// TIA Portal project "GzyHzy_1500" (V15)

(* hardware
DEVICE "S71500/ET200MP station_1"  S7-1500 station
   slot 0: "导轨_0"  Rack  6ES7 590-1***0-0AA0
   slot 0: "PM 70W 120/230VAC"  PM 70W 120/230VAC  6EP1332-4BA00
   slot 1: "1#DCC"  CPU 1511-1 PN  6ES7 511-1AK02-0AB0  V2.5
      slot 3: "CPU 显示_1"  6ES7591-1AA00-0AA0
   slot 2: "CP 1542-5_1"  CP 1542-5  6GK7 542-5FX00-0XE0  V1.0
   slot 3: "DI 32x24VDC BA_1"  DI 32x24VDC BA  6ES7 521-1BL10-0AA0  V1.0
   slot 4: "DQ 32x24VDC/0.5A BA_1"  DQ 32x24VDC/0.5A BA  6ES7 522-1BL10-0AA0  V1.0
   slot 5: "AI 8xU/I/RTD/TC ST_1"  AI 8xU/I/RTD/TC ST  6ES7 531-7KF00-0AB0  V2.1
   slot 6: "AI 8xU/I/RTD/TC ST_2"  AI 8xU/I/RTD/TC ST  6ES7 531-7KF00-0AB0  V2.1
   slot 7: "AI 8xU/I/RTD/TC ST_3"  AI 8xU/I/RTD/TC ST  6ES7 531-7KF00-0AB0  V2.1
   slot 8: "AI 8xU/I/RTD/TC ST_4"  AI 8xU/I/RTD/TC ST  6ES7 531-7KF00-0AB0  V2.1
   slot 9: "AI 8xU/I/RTD/TC ST_5"  AI 8xU/I/RTD/TC ST  6ES7 531-7KF00-0AB0  V2.1
   slot 10: "AQ 8xU/I HS_1"  AQ 8xU/I HS  6ES7 532-5HF00-0AB0  V2.1
DEVICE "GSD device_1"  GSD.Device
   slot 0: "机架_0"  Rail
   slot 0: "1#DCC_485"  PB-B-MODBUS  V2.0
DEVICE "S71500/ET200MP station_2"  S7-1500 station
   slot 0: "导轨_0"  Rack  6ES7 590-1***0-0AA0
   slot 0: "PM 70W 120/230VAC"  PM 70W 120/230VAC  6EP1332-4BA00
   slot 1: "1#GZY"  CPU 1511-1 PN  6ES7 511-1AK02-0AB0  V2.5
      slot 3: "CPU 显示_1"  6ES7591-1AA00-0AA0
   slot 2: "CP 1542-5_1"  CP 1542-5  6GK7 542-5FX00-0XE0  V1.0
   slot 3: "DI 32x24VDC BA_1"  DI 32x24VDC BA  6ES7 521-1BL10-0AA0  V1.0
   slot 4: "DI 32x24VDC BA_2"  DI 32x24VDC BA  6ES7 521-1BL10-0AA0  V1.0
   slot 5: "DI 32x24VDC BA_3"  DI 32x24VDC BA  6ES7 521-1BL10-0AA0  V1.0
   slot 6: "DQ 32x24VDC/0.5A BA_1"  DQ 32x24VDC/0.5A BA  6ES7 522-1BL10-0AA0  V1.0
   slot 7: "AI 8xU/I/RTD/TC ST_1"  AI 8xU/I/RTD/TC ST  6ES7 531-7KF00-0AB0  V2.1
   slot 8: "AI 8xU/I/RTD/TC ST_2"  AI 8xU/I/RTD/TC ST  6ES7 531-7KF00-0AB0  V2.1
   slot 9: "AI 8xU/I/RTD/TC ST_3"  AI 8xU/I/RTD/TC ST  6ES7 531-7KF00-0AB0  V2.1
   slot 10: "AI 8xU/I/RTD/TC ST_4"  AI 8xU/I/RTD/TC ST  6ES7 531-7KF00-0AB0  V2.1
   slot 11: "AQ 8xU/I HS_1"  AQ 8xU/I HS  6ES7 532-5HF00-0AB0  V2.1
DEVICE "S71500/ET200MP station_3"  S7-1500 station
   slot 0: "导轨_0"  Rack  6ES7 590-1***0-0AA0
   slot 0: "PM 70W 120/230VAC"  PM 70W 120/230VAC  6EP1332-4BA00
   slot 1: "1#HZY"  CPU 1511-1 PN  6ES7 511-1AK02-0AB0  V2.5
      slot 3: "CPU 显示_1"  6ES7591-1AA00-0AA0
   slot 2: "CP 1542-5_1"  CP 1542-5  6GK7 542-5FX00-0XE0  V1.0
   slot 3: "DI 32x24VDC BA_1"  DI 32x24VDC BA  6ES7 521-1BL10-0AA0  V1.0
   slot 4: "DI 32x24VDC BA_2"  DI 32x24VDC BA  6ES7 521-1BL10-0AA0  V1.0
   slot 5: "DQ 32x24VDC/0.5A BA_1"  DQ 32x24VDC/0.5A BA  6ES7 522-1BL10-0AA0  V1.0
   slot 6: "AI 8xU/I/RTD/TC ST_1"  AI 8xU/I/RTD/TC ST  6ES7 531-7KF00-0AB0  V2.1
   slot 7: "AI 8xU/I/RTD/TC ST_2"  AI 8xU/I/RTD/TC ST  6ES7 531-7KF00-0AB0  V2.1
   slot 8: "AQ 8xU/I HS_1"  AQ 8xU/I HS  6ES7 532-5HF00-0AB0  V2.1
DEVICE "S71500/ET200MP station_4"  S7-1500 station
   slot 0: "导轨_0"  Rack  6ES7 590-1***0-0AA0
   slot 2: "1#HZY_YTZ"  IM 155-5 DP ST  6ES7 155-5BA00-0AB0  V3.0
   slot 3: "DI 16x24VDC BA_1"  DI 16x24VDC BA  6ES7 521-1BH10-0AA0  V1.0
   slot 4: "DI 16x24VDC BA_2"  DI 16x24VDC BA  6ES7 521-1BH10-0AA0  V1.0
   slot 5: "DQ 16x24VDC/0.5A BA_1"  DQ 16x24VDC/0.5A BA  6ES7 522-1BH10-0AA0  V1.0
   slot 6: "AI 8xU/I/RTD/TC ST_1"  AI 8xU/I/RTD/TC ST  6ES7 531-7KF00-0AB0  V2.1
   slot 7: "AI 8xU/I/RTD/TC ST_2"  AI 8xU/I/RTD/TC ST  6ES7 531-7KF00-0AB0  V2.1
   slot 8: "AI 8xU/I/RTD/TC ST_3"  AI 8xU/I/RTD/TC ST  6ES7 531-7KF00-0AB0  V2.1
   slot 9: "AQ 8xU/I HS_1"  AQ 8xU/I HS  6ES7 532-5HF00-0AB0  V2.1
   slot 10: "DI 32x24VDC BA_1"  DI 32x24VDC BA  6ES7 521-1BL10-0AA0  V1.0
   slot 11: "AI 8xU/I/RTD/TC ST_4"  AI 8xU/I/RTD/TC ST  6ES7 531-7KF00-0AB0  V2.1
   slot 12: "AQ 8xU/I HS_2"  AQ 8xU/I HS  6ES7 532-5HF00-0AB0  V2.1
DEVICE "S71500/ET200MP station_5"  S7-1500 station
   slot 0: "导轨_0"  Rack  6ES7 590-1***0-0AA0
   slot 2: "1#HZY_PLZ"  IM 155-5 DP ST  6ES7 155-5BA00-0AB0  V3.0
   slot 3: "DI 16x24VDC BA_1"  DI 16x24VDC BA  6ES7 521-1BH10-0AA0  V1.0
   slot 4: "DI 16x24VDC BA_2"  DI 16x24VDC BA  6ES7 521-1BH10-0AA0  V1.0
   slot 5: "DI 16x24VDC BA_3"  DI 16x24VDC BA  6ES7 521-1BH10-0AA0  V1.0
   slot 6: "DQ 16x24VDC/0.5A BA_1"  DQ 16x24VDC/0.5A BA  6ES7 522-1BH10-0AA0  V1.0
   slot 7: "AI 8xU/I/RTD/TC ST_3"  AI 8xU/I/RTD/TC ST  6ES7 531-7KF00-0AB0  V2.1
   slot 8: "AQ 8xU/I HS_1"  AQ 8xU/I HS  6ES7 532-5HF00-0AB0  V2.1
DEVICE "GSD device_2"  GSD.Device
   slot 0: "机架_0"  Rail
   slot 0: "1#HZY_485"  PB-B-MODBUS  V2.0
DEVICE "GSD device_5"  GSD.Device
   slot 0: "机架_0"  Rail
   slot 0: "1#GZY_485"  PB-B-MODBUS  V2.0
DEVICE "S71500/ET200MP station_6"  S7-1500 station
   slot 0: "导轨_0"  Rack  6ES7 590-1***0-0AA0
   slot 0: "PM 70W 120/230VAC"  PM 70W 120/230VAC  6EP1332-4BA00
   slot 1: "2#DCC"  CPU 1511-1 PN  6ES7 511-1AK02-0AB0  V2.5
      slot 3: "CPU 显示_1"  6ES7591-1AA00-0AA0
   slot 2: "CP 1542-5_1"  CP 1542-5  6GK7 542-5FX00-0XE0  V1.0
   slot 3: "DI 32x24VDC BA_1"  DI 32x24VDC BA  6ES7 521-1BL10-0AA0  V1.0
   slot 4: "DQ 32x24VDC/0.5A BA_1"  DQ 32x24VDC/0.5A BA  6ES7 522-1BL10-0AA0  V1.0
   slot 5: "AI 8xU/I/RTD/TC ST_1"  AI 8xU/I/RTD/TC ST  6ES7 531-7KF00-0AB0  V2.1
   slot 6: "AI 8xU/I/RTD/TC ST_2"  AI 8xU/I/RTD/TC ST  6ES7 531-7KF00-0AB0  V2.1
   slot 7: "AI 8xU/I/RTD/TC ST_3"  AI 8xU/I/RTD/TC ST  6ES7 531-7KF00-0AB0  V2.1
   slot 8: "AI 8xU/I/RTD/TC ST_4"  AI 8xU/I/RTD/TC ST  6ES7 531-7KF00-0AB0  V2.1
   slot 9: "AI 8xU/I/RTD/TC ST_5"  AI 8xU/I/RTD/TC ST  6ES7 531-7KF00-0AB0  V2.1
   slot 10: "AQ 8xU/I HS_1"  AQ 8xU/I HS  6ES7 532-5HF00-0AB0  V2.1
DEVICE "GSD device_6"  GSD.Device
   slot 0: "机架_0"  Rail
   slot 0: "2#DCC_485"  PB-B-MODBUS  V2.0
DEVICE "S71500/ET200MP station_7"  S7-1500 station
   slot 0: "导轨_0"  Rack  6ES7 590-1***0-0AA0
   slot 0: "PM 70W 120/230VAC"  PM 70W 120/230VAC  6EP1332-4BA00
   slot 1: "2#GZY"  CPU 1511-1 PN  6ES7 511-1AK02-0AB0  V2.5
      slot 3: "CPU 显示_1"  6ES7591-1AA00-0AA0
   slot 2: "CP 1542-5_1"  CP 1542-5  6GK7 542-5FX00-0XE0  V1.0
   slot 3: "DI 32x24VDC BA_1"  DI 32x24VDC BA  6ES7 521-1BL10-0AA0  V1.0
   slot 4: "DI 32x24VDC BA_2"  DI 32x24VDC BA  6ES7 521-1BL10-0AA0  V1.0
   slot 5: "DI 32x24VDC BA_3"  DI 32x24VDC BA  6ES7 521-1BL10-0AA0  V1.0
   slot 6: "DQ 32x24VDC/0.5A BA_1"  DQ 32x24VDC/0.5A BA  6ES7 522-1BL10-0AA0  V1.0
   slot 7: "AI 8xU/I/RTD/TC ST_1"  AI 8xU/I/RTD/TC ST  6ES7 531-7KF00-0AB0  V2.1
   slot 8: "AI 8xU/I/RTD/TC ST_2"  AI 8xU/I/RTD/TC ST  6ES7 531-7KF00-0AB0  V2.1
   slot 9: "AI 8xU/I/RTD/TC ST_3"  AI 8xU/I/RTD/TC ST  6ES7 531-7KF00-0AB0  V2.1
   slot 10: "AI 8xU/I/RTD/TC ST_4"  AI 8xU/I/RTD/TC ST  6ES7 531-7KF00-0AB0  V2.1
   slot 11: "AQ 8xU/I HS_1"  AQ 8xU/I HS  6ES7 532-5HF00-0AB0  V2.1
DEVICE "GSD device_7"  GSD.Device
   slot 0: "机架_0"  Rail
   slot 0: "2#GZY_485"  PB-B-MODBUS  V2.0
DEVICE "S71500/ET200MP station_8"  S7-1500 station
   slot 0: "导轨_0"  Rack  6ES7 590-1***0-0AA0
   slot 0: "PM 70W 120/230VAC"  PM 70W 120/230VAC  6EP1332-4BA00
   slot 1: "2#HZY"  CPU 1511-1 PN  6ES7 511-1AK02-0AB0  V2.5
      slot 3: "CPU 显示_1"  6ES7591-1AA00-0AA0
   slot 2: "CP 1542-5_1"  CP 1542-5  6GK7 542-5FX00-0XE0  V1.0
   slot 3: "DI 32x24VDC BA_1"  DI 32x24VDC BA  6ES7 521-1BL10-0AA0  V1.0
   slot 4: "DI 32x24VDC BA_2"  DI 32x24VDC BA  6ES7 521-1BL10-0AA0  V1.0
   slot 5: "DQ 32x24VDC/0.5A BA_1"  DQ 32x24VDC/0.5A BA  6ES7 522-1BL10-0AA0  V1.0
   slot 6: "AI 8xU/I/RTD/TC ST_1"  AI 8xU/I/RTD/TC ST  6ES7 531-7KF00-0AB0  V2.1
   slot 7: "AI 8xU/I/RTD/TC ST_2"  AI 8xU/I/RTD/TC ST  6ES7 531-7KF00-0AB0  V2.1
   slot 8: "AQ 8xU/I HS_1"  AQ 8xU/I HS  6ES7 532-5HF00-0AB0  V2.1
DEVICE "S71500/ET200MP station_9"  S7-1500 station
   slot 0: "导轨_0"  Rack  6ES7 590-1***0-0AA0
   slot 2: "2#HZY_YTZ"  IM 155-5 DP ST  6ES7 155-5BA00-0AB0  V3.0
   slot 3: "DI 16x24VDC BA_1"  DI 16x24VDC BA  6ES7 521-1BH10-0AA0  V1.0
   slot 4: "DI 16x24VDC BA_2"  DI 16x24VDC BA  6ES7 521-1BH10-0AA0  V1.0
   slot 5: "DQ 16x24VDC/0.5A BA_1"  DQ 16x24VDC/0.5A BA  6ES7 522-1BH10-0AA0  V1.0
   slot 6: "AI 8xU/I/RTD/TC ST_1"  AI 8xU/I/RTD/TC ST  6ES7 531-7KF00-0AB0  V2.1
   slot 7: "AI 8xU/I/RTD/TC ST_2"  AI 8xU/I/RTD/TC ST  6ES7 531-7KF00-0AB0  V2.1
   slot 8: "AI 8xU/I/RTD/TC ST_3"  AI 8xU/I/RTD/TC ST  6ES7 531-7KF00-0AB0  V2.1
   slot 9: "AQ 8xU/I HS_1"  AQ 8xU/I HS  6ES7 532-5HF00-0AB0  V2.1
   slot 10: "DI 32x24VDC BA_1"  DI 32x24VDC BA  6ES7 521-1BL10-0AA0  V1.0
   slot 11: "AI 8xU/I/RTD/TC ST_4"  AI 8xU/I/RTD/TC ST  6ES7 531-7KF00-0AB0  V2.1
   slot 12: "AQ 8xU/I HS_2"  AQ 8xU/I HS  6ES7 532-5HF00-0AB0  V2.1
DEVICE "S71500/ET200MP station_10"  S7-1500 station
   slot 0: "导轨_0"  Rack  6ES7 590-1***0-0AA0
   slot 2: "2#HZY_PLZ"  IM 155-5 DP ST  6ES7 155-5BA00-0AB0  V3.0
   slot 3: "DI 16x24VDC BA_1"  DI 16x24VDC BA  6ES7 521-1BH10-0AA0  V1.0
   slot 4: "DI 16x24VDC BA_2"  DI 16x24VDC BA  6ES7 521-1BH10-0AA0  V1.0
   slot 5: "DI 16x24VDC BA_3"  DI 16x24VDC BA  6ES7 521-1BH10-0AA0  V1.0
   slot 6: "DQ 16x24VDC/0.5A BA_1"  DQ 16x24VDC/0.5A BA  6ES7 522-1BH10-0AA0  V1.0
   slot 7: "AI 8xU/I/RTD/TC ST_3"  AI 8xU/I/RTD/TC ST  6ES7 531-7KF00-0AB0  V2.1
   slot 8: "AQ 8xU/I HS_1"  AQ 8xU/I HS  6ES7 532-5HF00-0AB0  V2.1
DEVICE "GSD device_8"  GSD.Device
   slot 0: "机架_0"  Rail
   slot 0: "2#HZY_485"  PB-B-MODBUS  V2.0
DEVICE "S71500/ET200MP station_11"  S7-1500 station
   slot 0: "导轨_0"  Rack  6ES7 590-1***0-0AA0
   slot 0: "PM 70W 120/230VAC"  PM 70W 120/230VAC  6EP1332-4BA00
   slot 1: "3#GZY"  CPU 1511-1 PN  6ES7 511-1AK02-0AB0  V2.5
      slot 3: "CPU 显示_1"  6ES7591-1AA00-0AA0
   slot 2: "CP 1542-5_1"  CP 1542-5  6GK7 542-5FX00-0XE0  V1.0
   slot 3: "DI 32x24VDC BA_1"  DI 32x24VDC BA  6ES7 521-1BL10-0AA0  V1.0
   slot 4: "DI 32x24VDC BA_2"  DI 32x24VDC BA  6ES7 521-1BL10-0AA0  V1.0
   slot 5: "DI 32x24VDC BA_3"  DI 32x24VDC BA  6ES7 521-1BL10-0AA0  V1.0
   slot 6: "DQ 32x24VDC/0.5A BA_1"  DQ 32x24VDC/0.5A BA  6ES7 522-1BL10-0AA0  V1.0
   slot 7: "AI 8xU/I/RTD/TC ST_1"  AI 8xU/I/RTD/TC ST  6ES7 531-7KF00-0AB0  V2.1
   slot 8: "AI 8xU/I/RTD/TC ST_2"  AI 8xU/I/RTD/TC ST  6ES7 531-7KF00-0AB0  V2.1
   slot 9: "AI 8xU/I/RTD/TC ST_3"  AI 8xU/I/RTD/TC ST  6ES7 531-7KF00-0AB0  V2.1
   slot 10: "AI 8xU/I/RTD/TC ST_4"  AI 8xU/I/RTD/TC ST  6ES7 531-7KF00-0AB0  V2.1
   slot 11: "AQ 8xU/I HS_1"  AQ 8xU/I HS  6ES7 532-5HF00-0AB0  V2.1
DEVICE "GSD device_11"  GSD.Device
   slot 0: "机架_0"  Rail
   slot 0: "3#GZY_485"  PB-B-MODBUS  V2.0
DEVICE "S71500/ET200MP station_12"  S7-1500 station
   slot 0: "导轨_0"  Rack  6ES7 590-1***0-0AA0
   slot 0: "PM 70W 120/230VAC"  PM 70W 120/230VAC  6EP1332-4BA00
   slot 1: "3#HZY"  CPU 1511-1 PN  6ES7 511-1AK02-0AB0  V2.5
      slot 3: "CPU 显示_1"  6ES7591-1AA00-0AA0
   slot 2: "CP 1542-5_1"  CP 1542-5  6GK7 542-5FX00-0XE0  V1.0
   slot 3: "DI 32x24VDC BA_1"  DI 32x24VDC BA  6ES7 521-1BL10-0AA0  V1.0
   slot 4: "DI 32x24VDC BA_2"  DI 32x24VDC BA  6ES7 521-1BL10-0AA0  V1.0
   slot 5: "DQ 32x24VDC/0.5A BA_1"  DQ 32x24VDC/0.5A BA  6ES7 522-1BL10-0AA0  V1.0
   slot 6: "AI 8xU/I/RTD/TC ST_1"  AI 8xU/I/RTD/TC ST  6ES7 531-7KF00-0AB0  V2.1
   slot 7: "AI 8xU/I/RTD/TC ST_2"  AI 8xU/I/RTD/TC ST  6ES7 531-7KF00-0AB0  V2.1
   slot 8: "AQ 8xU/I HS_1"  AQ 8xU/I HS  6ES7 532-5HF00-0AB0  V2.1
DEVICE "S71500/ET200MP station_14"  S7-1500 station
   slot 0: "导轨_0"  Rack  6ES7 590-1***0-0AA0
   slot 2: "3#HZY_YTZ"  IM 155-5 DP ST  6ES7 155-5BA00-0AB0  V3.0
   slot 3: "DI 16x24VDC BA_1"  DI 16x24VDC BA  6ES7 521-1BH10-0AA0  V1.0
   slot 4: "DI 16x24VDC BA_2"  DI 16x24VDC BA  6ES7 521-1BH10-0AA0  V1.0
   slot 5: "DQ 16x24VDC/0.5A BA_1"  DQ 16x24VDC/0.5A BA  6ES7 522-1BH10-0AA0  V1.0
   slot 6: "AI 8xU/I/RTD/TC ST_1"  AI 8xU/I/RTD/TC ST  6ES7 531-7KF00-0AB0  V2.1
   slot 7: "AI 8xU/I/RTD/TC ST_2"  AI 8xU/I/RTD/TC ST  6ES7 531-7KF00-0AB0  V2.1
   slot 8: "AI 8xU/I/RTD/TC ST_3"  AI 8xU/I/RTD/TC ST  6ES7 531-7KF00-0AB0  V2.1
   slot 9: "AQ 8xU/I HS_1"  AQ 8xU/I HS  6ES7 532-5HF00-0AB0  V2.1
   slot 10: "DI 32x24VDC BA_1"  DI 32x24VDC BA  6ES7 521-1BL10-0AA0  V1.0
   slot 11: "AI 8xU/I/RTD/TC ST_4"  AI 8xU/I/RTD/TC ST  6ES7 531-7KF00-0AB0  V2.1
   slot 12: "AQ 8xU/I HS_2"  AQ 8xU/I HS  6ES7 532-5HF00-0AB0  V2.1
DEVICE "S71500/ET200MP station_13"  S7-1500 station
   slot 0: "导轨_0"  Rack  6ES7 590-1***0-0AA0
   slot 2: "3#HZY_PLZ"  IM 155-5 DP ST  6ES7 155-5BA00-0AB0  V3.0
   slot 3: "DI 16x24VDC BA_1"  DI 16x24VDC BA  6ES7 521-1BH10-0AA0  V1.0
   slot 4: "DI 16x24VDC BA_2"  DI 16x24VDC BA  6ES7 521-1BH10-0AA0  V1.0
   slot 5: "DI 16x24VDC BA_3"  DI 16x24VDC BA  6ES7 521-1BH10-0AA0  V1.0
   slot 6: "DQ 16x24VDC/0.5A BA_1"  DQ 16x24VDC/0.5A BA  6ES7 522-1BH10-0AA0  V1.0
   slot 7: "AI 8xU/I/RTD/TC ST_3"  AI 8xU/I/RTD/TC ST  6ES7 531-7KF00-0AB0  V2.1
   slot 8: "AQ 8xU/I HS_1"  AQ 8xU/I HS  6ES7 532-5HF00-0AB0  V2.1
DEVICE "GSD device_12"  GSD.Device
   slot 0: "机架_0"  Rail
   slot 0: "3#HZY_485"  PB-B-MODBUS  V2.0
DEVICE "S71500/ET200MP station_15"  S7-1500 station
   slot 0: "导轨_0"  Rack  6ES7 590-1***0-0AA0
   slot 0: "PM 70W 120/230VAC"  PM 70W 120/230VAC  6EP1332-4BA00
   slot 1: "4#GZY"  CPU 1511-1 PN  6ES7 511-1AK02-0AB0  V2.5
      slot 3: "CPU 显示_1"  6ES7591-1AA00-0AA0
   slot 2: "CP 1542-5_1"  CP 1542-5  6GK7 542-5FX00-0XE0  V1.0
   slot 3: "DI 32x24VDC BA_1"  DI 32x24VDC BA  6ES7 521-1BL10-0AA0  V1.0
   slot 4: "DI 32x24VDC BA_2"  DI 32x24VDC BA  6ES7 521-1BL10-0AA0  V1.0
   slot 5: "DI 32x24VDC BA_3"  DI 32x24VDC BA  6ES7 521-1BL10-0AA0  V1.0
   slot 6: "DQ 32x24VDC/0.5A BA_1"  DQ 32x24VDC/0.5A BA  6ES7 522-1BL10-0AA0  V1.0
   slot 7: "AI 8xU/I/RTD/TC ST_1"  AI 8xU/I/RTD/TC ST  6ES7 531-7KF00-0AB0  V2.1
   slot 8: "AI 8xU/I/RTD/TC ST_2"  AI 8xU/I/RTD/TC ST  6ES7 531-7KF00-0AB0  V2.1
   slot 9: "AI 8xU/I/RTD/TC ST_3"  AI 8xU/I/RTD/TC ST  6ES7 531-7KF00-0AB0  V2.1
   slot 10: "AI 8xU/I/RTD/TC ST_4"  AI 8xU/I/RTD/TC ST  6ES7 531-7KF00-0AB0  V2.1
   slot 11: "AQ 8xU/I HS_1"  AQ 8xU/I HS  6ES7 532-5HF00-0AB0  V2.1
DEVICE "S71500/ET200MP station_16"  S7-1500 station
   slot 0: "导轨_0"  Rack  6ES7 590-1***0-0AA0
   slot 0: "PM 70W 120/230VAC"  PM 70W 120/230VAC  6EP1332-4BA00
   slot 1: "4#HZY"  CPU 1511-1 PN  6ES7 511-1AK02-0AB0  V2.5
      slot 3: "CPU 显示_1"  6ES7591-1AA00-0AA0
   slot 2: "CP 1542-5_1"  CP 1542-5  6GK7 542-5FX00-0XE0  V1.0
   slot 3: "DI 32x24VDC BA_1"  DI 32x24VDC BA  6ES7 521-1BL10-0AA0  V1.0
   slot 4: "DI 32x24VDC BA_2"  DI 32x24VDC BA  6ES7 521-1BL10-0AA0  V1.0
   slot 5: "DQ 32x24VDC/0.5A BA_1"  DQ 32x24VDC/0.5A BA  6ES7 522-1BL10-0AA0  V1.0
   slot 6: "AI 8xU/I/RTD/TC ST_1"  AI 8xU/I/RTD/TC ST  6ES7 531-7KF00-0AB0  V2.1
   slot 7: "AI 8xU/I/RTD/TC ST_2"  AI 8xU/I/RTD/TC ST  6ES7 531-7KF00-0AB0  V2.1
   slot 8: "AQ 8xU/I HS_1"  AQ 8xU/I HS  6ES7 532-5HF00-0AB0  V2.1
DEVICE "S71500/ET200MP station_17"  S7-1500 station
   slot 0: "导轨_0"  Rack  6ES7 590-1***0-0AA0
   slot 2: "4#HZY_YTZ"  IM 155-5 DP ST  6ES7 155-5BA00-0AB0  V3.0
   slot 3: "DI 16x24VDC BA_1"  DI 16x24VDC BA  6ES7 521-1BH10-0AA0  V1.0
   slot 4: "DI 16x24VDC BA_2"  DI 16x24VDC BA  6ES7 521-1BH10-0AA0  V1.0
   slot 5: "DQ 16x24VDC/0.5A BA_1"  DQ 16x24VDC/0.5A BA  6ES7 522-1BH10-0AA0  V1.0
   slot 6: "AI 8xU/I/RTD/TC ST_1"  AI 8xU/I/RTD/TC ST  6ES7 531-7KF00-0AB0  V2.1
   slot 7: "AI 8xU/I/RTD/TC ST_2"  AI 8xU/I/RTD/TC ST  6ES7 531-7KF00-0AB0  V2.1
   slot 8: "AI 8xU/I/RTD/TC ST_3"  AI 8xU/I/RTD/TC ST  6ES7 531-7KF00-0AB0  V2.1
   slot 9: "AQ 8xU/I HS_1"  AQ 8xU/I HS  6ES7 532-5HF00-0AB0  V2.1
   slot 10: "DI 32x24VDC BA_1"  DI 32x24VDC BA  6ES7 521-1BL10-0AA0  V1.0
   slot 11: "AI 8xU/I/RTD/TC ST_4"  AI 8xU/I/RTD/TC ST  6ES7 531-7KF00-0AB0  V2.1
   slot 12: "AQ 8xU/I HS_2"  AQ 8xU/I HS  6ES7 532-5HF00-0AB0  V2.1
DEVICE "S71500/ET200MP station_18"  S7-1500 station
   slot 0: "导轨_0"  Rack  6ES7 590-1***0-0AA0
   slot 2: "4#HZY_PLZ"  IM 155-5 DP ST  6ES7 155-5BA00-0AB0  V3.0
   slot 3: "DI 16x24VDC BA_1"  DI 16x24VDC BA  6ES7 521-1BH10-0AA0  V1.0
   slot 4: "DI 16x24VDC BA_2"  DI 16x24VDC BA  6ES7 521-1BH10-0AA0  V1.0
   slot 5: "DI 16x24VDC BA_3"  DI 16x24VDC BA  6ES7 521-1BH10-0AA0  V1.0
   slot 6: "DQ 16x24VDC/0.5A BA_1"  DQ 16x24VDC/0.5A BA  6ES7 522-1BH10-0AA0  V1.0
   slot 7: "AI 8xU/I/RTD/TC ST_3"  AI 8xU/I/RTD/TC ST  6ES7 531-7KF00-0AB0  V2.1
   slot 8: "AQ 8xU/I HS_1"  AQ 8xU/I HS  6ES7 532-5HF00-0AB0  V2.1
DEVICE "GSD device_16"  GSD.Device
   slot 0: "机架_0"  Rail
   slot 0: "4#HZY_485"  PB-B-MODBUS  V2.0
DEVICE "S71500/ET200MP station_19"  S7-1500 station
   slot 0: "导轨_0"  Rack  6ES7 590-1***0-0AA0
   slot 0: "PM 70W 120/230VAC"  PM 70W 120/230VAC  6EP1332-4BA00
   slot 1: "1#LM"  CPU 1511-1 PN  6ES7 511-1AK02-0AB0  V2.5
      slot 3: "CPU 显示_1"  6ES7591-1AA00-0AA0
   slot 2: "CP 1542-5_1"  CP 1542-5  6GK7 542-5FX00-0XE0  V1.0
   slot 3: "DI 32x24VDC BA_1"  DI 32x24VDC BA  6ES7 521-1BL10-0AA0  V1.0
   slot 4: "DI 32x24VDC BA_2"  DI 32x24VDC BA  6ES7 521-1BL10-0AA0  V1.0
   slot 5: "DI 32x24VDC BA_3"  DI 32x24VDC BA  6ES7 521-1BL10-0AA0  V1.0
   slot 6: "DQ 32x24VDC/0.5A BA_1"  DQ 32x24VDC/0.5A BA  6ES7 522-1BL10-0AA0  V1.0
   slot 7: "AI 8xU/I/RTD/TC ST_1"  AI 8xU/I/RTD/TC ST  6ES7 531-7KF00-0AB0  V2.1
   slot 8: "AI 8xU/I/RTD/TC ST_2"  AI 8xU/I/RTD/TC ST  6ES7 531-7KF00-0AB0  V2.1
   slot 9: "AI 8xU/I/RTD/TC ST_3"  AI 8xU/I/RTD/TC ST  6ES7 531-7KF00-0AB0  V2.1
   slot 10: "AQ 8xU/I HS_1"  AQ 8xU/I HS  6ES7 532-5HF00-0AB0  V2.1
DEVICE "GSD device_19"  GSD.Device
   slot 0: "机架_0"  Rail
   slot 0: "1#LM_485"  PB-B-MODBUS  V2.0
DEVICE "GSD device_15"  GSD.Device
   slot 0: "机架_0"  Rail
   slot 0: "4#GZY_485"  PB-B-MODBUS  V2.0
DEVICE "GSD device_28"  GSD.Device
   slot 0: "机架_0"  Rail
DEVICE "GSD device_25"  GSD.Device
   slot 0: "机架_0"  Rail
DEVICE "GSD device_21"  GSD.Device
   slot 0: "机架_0"  Rail
DEVICE "GSD device_22"  GSD.Device
   slot 0: "机架_0"  Rail
DEVICE "SINAMICS G_4"  Sinamics.Device
   slot 0: "	_0"  Rail  SinamicsG120Rack-V
   slot 2: "电炉料罐车变频_1"  G120 CU240E-2  6SL3244-0BB12-1BA1  4.7.6
   slot 3: "PM240-2 IP20"  PM240-2 IP20  6SL3210-1PE23-3ULx  -
DEVICE "GSD device_23"  GSD.Device
   slot 0: "机架_0"  Rail
DEVICE "GSD device_24"  GSD.Device
   slot 0: "机架_0"  Rail
DEVICE "GSD device_26"  GSD.Device
   slot 0: "机架_0"  Rail
DEVICE "GSD device_3"  GSD.Device
   slot 0: "机架_0"  Rail
DEVICE "GSD device_4"  GSD.Device
   slot 0: "机架_0"  Rail
DEVICE "GSD device_9"  GSD.Device
   slot 0: "机架_0"  Rail
DEVICE "GSD device_10"  GSD.Device
   slot 0: "机架_0"  Rail
DEVICE "GSD device_13"  GSD.Device
   slot 0: "机架_0"  Rail
DEVICE "GSD device_14"  GSD.Device
   slot 0: "机架_0"  Rail
DEVICE "GSD device_17"  GSD.Device
   slot 0: "机架_0"  Rail
DEVICE "GSD device_18"  GSD.Device
   slot 0: "机架_0"  Rail
DEVICE "S71500/ET200MP station_20"  S7-1500 station
   slot 0: "导轨_0"  Rack  6ES7 590-1***0-0AA0
   slot 0: "PM 70W 120/230VAC"  PM 70W 120/230VAC  6EP1332-4BA00
   slot 1: "1#SBF"  CPU 1511-1 PN  6ES7 511-1AK02-0AB0  V2.5
      slot 3: "CPU 显示_1"  6ES7591-1AA00-0AA0
   slot 2: "CP 1542-5_1"  CP 1542-5  6GK7 542-5FX00-0XE0  V1.0
   slot 3: "DI 32x24VDC BA_1"  DI 32x24VDC BA  6ES7 521-1BL10-0AA0  V1.0
   slot 4: "DI 32x24VDC BA_2"  DI 32x24VDC BA  6ES7 521-1BL10-0AA0  V1.0
   slot 5: "DI 32x24VDC BA_3"  DI 32x24VDC BA  6ES7 521-1BL10-0AA0  V1.0
   slot 6: "DI 32x24VDC BA_4"  DI 32x24VDC BA  6ES7 521-1BL10-0AA0  V1.0
   slot 7: "DI 32x24VDC BA_5"  DI 32x24VDC BA  6ES7 521-1BL10-0AA0  V1.0
   slot 8: "DI 32x24VDC BA_6"  DI 32x24VDC BA  6ES7 521-1BL10-0AA0  V1.0
   slot 9: "PS 25W 24VDC_1"  PS 25W 24VDC  6ES7 505-0KA00-0AB0  V1.0
   slot 10: "DQ 32x24VDC/0.5A BA_1"  DQ 32x24VDC/0.5A BA  6ES7 522-1BL10-0AA0  V1.0
   slot 11: "DQ 32x24VDC/0.5A BA_2"  DQ 32x24VDC/0.5A BA  6ES7 522-1BL10-0AA0  V1.0
DEVICE "S71500/ET200MP station_25"  S7-1500 station
   slot 0: "导轨_0"  Rack  6ES7 590-1***0-0AA0
   slot 0: "PM 70W 120/230VAC"  PM 70W 120/230VAC  6EP1332-4BA00
   slot 1: "2#SBF"  CPU 1511-1 PN  6ES7 511-1AK02-0AB0  V2.5
      slot 3: "CPU 显示_1"  6ES7591-1AA00-0AA0
   slot 2: "CP 1542-5_1"  CP 1542-5  6GK7 542-5FX00-0XE0  V1.0
   slot 3: "DI 32x24VDC BA_1"  DI 32x24VDC BA  6ES7 521-1BL10-0AA0  V1.0
   slot 4: "DI 32x24VDC BA_2"  DI 32x24VDC BA  6ES7 521-1BL10-0AA0  V1.0
   slot 5: "DI 32x24VDC BA_3"  DI 32x24VDC BA  6ES7 521-1BL10-0AA0  V1.0
   slot 6: "DI 32x24VDC BA_4"  DI 32x24VDC BA  6ES7 521-1BL10-0AA0  V1.0
   slot 7: "DI 32x24VDC BA_5"  DI 32x24VDC BA  6ES7 521-1BL10-0AA0  V1.0
   slot 8: "DI 32x24VDC BA_6"  DI 32x24VDC BA  6ES7 521-1BL10-0AA0  V1.0
   slot 9: "PS 25W 24VDC_1"  PS 25W 24VDC  6ES7 505-0KA00-0AB0  V1.0
   slot 10: "DQ 32x24VDC/0.5A BA_1"  DQ 32x24VDC/0.5A BA  6ES7 522-1BL10-0AA0  V1.0
   slot 11: "DQ 32x24VDC/0.5A BA_2"  DQ 32x24VDC/0.5A BA  6ES7 522-1BL10-0AA0  V1.0
DEVICE "S71500/ET200MP station_21"  S7-1500 station
   slot 0: "导轨_0"  Rack  6ES7 590-1***0-0AA0
   slot 2: "1#SBF_1"  IM 155-5 DP ST  6ES7 155-5BA00-0AB0  V3.0
   slot 3: "DI 32x24VDC BA_1"  DI 32x24VDC BA  6ES7 521-1BL10-0AA0  V1.0
   slot 4: "DI 32x24VDC BA_2"  DI 32x24VDC BA  6ES7 521-1BL10-0AA0  V1.0
   slot 5: "DI 32x24VDC BA_3"  DI 32x24VDC BA  6ES7 521-1BL10-0AA0  V1.0
   slot 6: "DQ 32x24VDC/0.5A BA_1"  DQ 32x24VDC/0.5A BA  6ES7 522-1BL10-0AA0  V1.0
   slot 7: "DQ 32x24VDC/0.5A BA_2"  DQ 32x24VDC/0.5A BA  6ES7 522-1BL10-0AA0  V1.0
DEVICE "S71500/ET200MP station_22"  S7-1500 station
   slot 0: "导轨_0"  Rack  6ES7 590-1***0-0AA0
   slot 2: "1#SBF_2"  IM 155-5 DP ST  6ES7 155-5BA00-0AB0  V3.0
   slot 3: "AI 8xU/I/RTD/TC ST_1"  AI 8xU/I/RTD/TC ST  6ES7 531-7KF00-0AB0  V2.1
   slot 4: "AI 8xU/I/RTD/TC ST_2"  AI 8xU/I/RTD/TC ST  6ES7 531-7KF00-0AB0  V2.1
   slot 5: "AI 8xU/I/RTD/TC ST_3"  AI 8xU/I/RTD/TC ST  6ES7 531-7KF00-0AB0  V2.1
   slot 6: "AI 8xU/I/RTD/TC ST_4"  AI 8xU/I/RTD/TC ST  6ES7 531-7KF00-0AB0  V2.1
   slot 7: "AI 8xU/I/RTD/TC ST_5"  AI 8xU/I/RTD/TC ST  6ES7 531-7KF00-0AB0  V2.1
   slot 8: "AQ 8xU/I HS_1"  AQ 8xU/I HS  6ES7 532-5HF00-0AB0  V2.1
   slot 9: "AQ 8xU/I HS_2"  AQ 8xU/I HS  6ES7 532-5HF00-0AB0  V2.1
   slot 10: "AQ 8xU/I HS_3"  AQ 8xU/I HS  6ES7 532-5HF00-0AB0  V2.1
DEVICE "S71500/ET200MP station_23"  S7-1500 station
   slot 0: "导轨_0"  Rack  6ES7 590-1***0-0AA0
   slot 2: "1#SBF_3"  IM 155-5 DP ST  6ES7 155-5BA00-0AB0  V3.0
   slot 3: "DI 32x24VDC BA_1"  DI 32x24VDC BA  6ES7 521-1BL10-0AA0  V1.0
   slot 4: "DI 32x24VDC BA_2"  DI 32x24VDC BA  6ES7 521-1BL10-0AA0  V1.0
   slot 5: "DQ 32x24VDC/0.5A BA_1"  DQ 32x24VDC/0.5A BA  6ES7 522-1BL10-0AA0  V1.0
   slot 6: "AI 8xU/I/RTD/TC ST_1"  AI 8xU/I/RTD/TC ST  6ES7 531-7KF00-0AB0  V2.1
   slot 7: "AI 8xU/I/RTD/TC ST_2"  AI 8xU/I/RTD/TC ST  6ES7 531-7KF00-0AB0  V2.1
   slot 8: "AQ 8xU/I HS_1"  AQ 8xU/I HS  6ES7 532-5HF00-0AB0  V2.1
DEVICE "S71500/ET200MP station_24"  S7-1500 station
   slot 0: "导轨_0"  Rack  6ES7 590-1***0-0AA0
   slot 2: "1#SBF_4"  IM 155-5 DP ST  6ES7 155-5BA00-0AB0  V3.0
   slot 3: "DI 32x24VDC BA_1"  DI 32x24VDC BA  6ES7 521-1BL10-0AA0  V1.0
   slot 4: "DI 32x24VDC BA_2"  DI 32x24VDC BA  6ES7 521-1BL10-0AA0  V1.0
   slot 5: "DQ 32x24VDC/0.5A BA_1"  DQ 32x24VDC/0.5A BA  6ES7 522-1BL10-0AA0  V1.0
   slot 6: "AI 8xU/I/RTD/TC ST_1"  AI 8xU/I/RTD/TC ST  6ES7 531-7KF00-0AB0  V2.1
   slot 7: "AI 8xU/I/RTD/TC ST_2"  AI 8xU/I/RTD/TC ST  6ES7 531-7KF00-0AB0  V2.1
   slot 8: "AQ 8xU/I HS_1"  AQ 8xU/I HS  6ES7 532-5HF00-0AB0  V2.1
DEVICE "S71500/ET200MP station_26"  S7-1500 station
   slot 0: "导轨_0"  Rack  6ES7 590-1***0-0AA0
   slot 2: "2#SBF_1"  IM 155-5 DP ST  6ES7 155-5BA00-0AB0  V3.0
   slot 3: "DI 32x24VDC BA_1"  DI 32x24VDC BA  6ES7 521-1BL10-0AA0  V1.0
   slot 4: "DI 32x24VDC BA_2"  DI 32x24VDC BA  6ES7 521-1BL10-0AA0  V1.0
   slot 5: "DI 32x24VDC BA_3"  DI 32x24VDC BA  6ES7 521-1BL10-0AA0  V1.0
   slot 6: "DQ 32x24VDC/0.5A BA_1"  DQ 32x24VDC/0.5A BA  6ES7 522-1BL10-0AA0  V1.0
   slot 7: "DQ 32x24VDC/0.5A BA_2"  DQ 32x24VDC/0.5A BA  6ES7 522-1BL10-0AA0  V1.0
DEVICE "S71500/ET200MP station_27"  S7-1500 station
   slot 0: "导轨_0"  Rack  6ES7 590-1***0-0AA0
   slot 2: "2#SBF_2"  IM 155-5 DP ST  6ES7 155-5BA00-0AB0  V3.0
   slot 3: "AI 8xU/I/RTD/TC ST_1"  AI 8xU/I/RTD/TC ST  6ES7 531-7KF00-0AB0  V2.1
   slot 4: "AI 8xU/I/RTD/TC ST_2"  AI 8xU/I/RTD/TC ST  6ES7 531-7KF00-0AB0  V2.1
   slot 5: "AI 8xU/I/RTD/TC ST_3"  AI 8xU/I/RTD/TC ST  6ES7 531-7KF00-0AB0  V2.1
   slot 6: "AI 8xU/I/RTD/TC ST_4"  AI 8xU/I/RTD/TC ST  6ES7 531-7KF00-0AB0  V2.1
   slot 7: "AI 8xU/I/RTD/TC ST_5"  AI 8xU/I/RTD/TC ST  6ES7 531-7KF00-0AB0  V2.1
   slot 8: "AQ 8xU/I HS_1"  AQ 8xU/I HS  6ES7 532-5HF00-0AB0  V2.1
   slot 9: "AQ 8xU/I HS_2"  AQ 8xU/I HS  6ES7 532-5HF00-0AB0  V2.1
   slot 10: "AQ 8xU/I HS_3"  AQ 8xU/I HS  6ES7 532-5HF00-0AB0  V2.1
DEVICE "S71500/ET200MP station_28"  S7-1500 station
   slot 0: "导轨_0"  Rack  6ES7 590-1***0-0AA0
   slot 2: "2#SBF_3"  IM 155-5 DP ST  6ES7 155-5BA00-0AB0  V3.0
   slot 3: "DI 32x24VDC BA_1"  DI 32x24VDC BA  6ES7 521-1BL10-0AA0  V1.0
   slot 4: "DI 32x24VDC BA_2"  DI 32x24VDC BA  6ES7 521-1BL10-0AA0  V1.0
   slot 5: "DQ 32x24VDC/0.5A BA_1"  DQ 32x24VDC/0.5A BA  6ES7 522-1BL10-0AA0  V1.0
   slot 6: "AI 8xU/I/RTD/TC ST_1"  AI 8xU/I/RTD/TC ST  6ES7 531-7KF00-0AB0  V2.1
   slot 7: "AI 8xU/I/RTD/TC ST_2"  AI 8xU/I/RTD/TC ST  6ES7 531-7KF00-0AB0  V2.1
   slot 8: "AQ 8xU/I HS_1"  AQ 8xU/I HS  6ES7 532-5HF00-0AB0  V2.1
DEVICE "S71500/ET200MP station_29"  S7-1500 station
   slot 0: "导轨_0"  Rack  6ES7 590-1***0-0AA0
   slot 2: "2#SBF_4"  IM 155-5 DP ST  6ES7 155-5BA00-0AB0  V3.0
   slot 3: "DI 32x24VDC BA_1"  DI 32x24VDC BA  6ES7 521-1BL10-0AA0  V1.0
   slot 4: "DI 32x24VDC BA_2"  DI 32x24VDC BA  6ES7 521-1BL10-0AA0  V1.0
   slot 5: "DQ 32x24VDC/0.5A BA_1"  DQ 32x24VDC/0.5A BA  6ES7 522-1BL10-0AA0  V1.0
   slot 6: "AI 8xU/I/RTD/TC ST_1"  AI 8xU/I/RTD/TC ST  6ES7 531-7KF00-0AB0  V2.1
   slot 7: "AI 8xU/I/RTD/TC ST_2"  AI 8xU/I/RTD/TC ST  6ES7 531-7KF00-0AB0  V2.1
   slot 8: "AQ 8xU/I HS_1"  AQ 8xU/I HS  6ES7 532-5HF00-0AB0  V2.1
DEVICE "S71500/ET200MP station_30"  S7-1500 station
   slot 0: "导轨_0"  Rack  6ES7 590-1***0-0AA0
   slot 0: "PM 70W 120/230VAC"  PM 70W 120/230VAC  6EP1332-4BA00
   slot 1: "2#LM"  CPU 1511-1 PN  6ES7 511-1AK02-0AB0  V2.5
      slot 3: "CPU 显示_1"  6ES7591-1AA00-0AA0
   slot 2: "CP 1542-5_1"  CP 1542-5  6GK7 542-5FX00-0XE0  V1.0
   slot 3: "DI 32x24VDC BA_1"  DI 32x24VDC BA  6ES7 521-1BL10-0AA0  V1.0
   slot 4: "DI 32x24VDC BA_2"  DI 32x24VDC BA  6ES7 521-1BL10-0AA0  V1.0
   slot 5: "DI 32x24VDC BA_3"  DI 32x24VDC BA  6ES7 521-1BL10-0AA0  V1.0
   slot 6: "DQ 32x24VDC/0.5A BA_1"  DQ 32x24VDC/0.5A BA  6ES7 522-1BL10-0AA0  V1.0
   slot 7: "AI 8xU/I/RTD/TC ST_1"  AI 8xU/I/RTD/TC ST  6ES7 531-7KF00-0AB0  V2.1
   slot 8: "AI 8xU/I/RTD/TC ST_2"  AI 8xU/I/RTD/TC ST  6ES7 531-7KF00-0AB0  V2.1
   slot 9: "AI 8xU/I/RTD/TC ST_3"  AI 8xU/I/RTD/TC ST  6ES7 531-7KF00-0AB0  V2.1
   slot 10: "AQ 8xU/I HS_1"  AQ 8xU/I HS  6ES7 532-5HF00-0AB0  V2.1
DEVICE "GSD device_27"  GSD.Device
   slot 0: "机架_0"  Rail
   slot 0: "2#LM_485"  PB-B-MODBUS  V2.0
DEVICE "GSD device_30"  GSD.Device
   slot 0: "机架_0"  Rail
DEVICE "GSD device_31"  GSD.Device
   slot 0: "机架_0"  Rail
DEVICE "GSD device_32"  GSD.Device
   slot 0: "机架_0"  Rail
*)

// ===== PLC "1#DCC"  CPU 1511-1 PN =====

VAR_GLOBAL   // PLC tag table "默认变量表"
   "2#2号电场一次运行电压" AT %IW296 : Int;
   "2#2号电场二次运行电压" AT %IW300 : Int;
   "2#1号电场就绪" AT %I2.1 : Bool;
   "2#除尘热风管进口温度" AT %IW332 : Int;
   "2#电场热风管入口压力" AT %IW324 : Int;
   "1#3号电场二次运行电流" AT %IW278 : Int;
   "1#3号电场一次运行电压" AT %IW272 : Int;
   "1#3号电场二次运行电压" AT %IW276 : Int;
   "2#2号电场备妥" AT %I2.4 : Bool;
   "2#1号电场故障" AT %I2.3 : Bool;
   "2#4号电场二次运行电流" AT %IW318 : Int;
   "1#电场热风管出口压力" AT %IW322 : Int;
   "1#除尘热风管进口温度" AT %IW328 : Int;
   "1#电场热风管入口压力" AT %IW320 : Int;
   "1#3号电场运行" AT %I1.2 : Bool;
   "1#除尘热风管出口温度" AT %IW330 : Int;
   "1#3号电场一次运行电流" AT %IW274 : Int;
   "2#1号电场备妥" AT %I2.0 : Bool;
   "2#3号电场二次运行电流" AT %IW310 : Int;
   "2#3号电场一次运行电压" AT %IW304 : Int;
   "2#2号电场运行" AT %I2.6 : Bool;
   "2#除尘热风管出口温度" AT %IW334 : Int;
   "2#电场热风管出口压力" AT %IW326 : Int;
   "2#4号电场一次运行电流" AT %IW314 : Int;
   "1#1号电场一次运行电流" AT %IW258 : Int;
   "1#2号电场一次运行电流" AT %IW266 : Int;
   "2#3号电场一次运行电流" AT %IW306 : Int;
   "2#2号电场一次运行电流" AT %IW298 : Int;
   "2#1号电场一次运行电流" AT %IW290 : Int;
   "1#4号电场一次运行电流" AT %IW282 : Int;
   "1#1号电场二次运行电流" AT %IW262 : Int;
   "1#1号电场一次运行电压" AT %IW256 : Int;
   "1#1号电场二次运行电压" AT %IW260 : Int;
   "1#1号电场运行" AT %I0.2 : Bool;
   "1#1号电场就绪" AT %I0.1 : Bool;
   "2#3号电场二次运行电压" AT %IW308 : Int;
   "1#2号电场二次运行电流" AT %IW270 : Int;
   "1#2号电场一次运行电压" AT %IW264 : Int;
   "1#3号电场备妥" AT %I1.0 : Bool;
   "1#2号电场故障" AT %I0.7 : Bool;
   "1#4号电场二次运行电流" AT %IW286 : Int;
   "1#4号电场运行" AT %I1.6 : Bool;
   "1#4号电场就绪" AT %I1.5 : Bool;
   "2#2号电场二次运行电流" AT %IW302 : Int;
   "2#4号电场一次运行电压" AT %IW312 : Int;
   "2#4号电场二次运行电压" AT %IW316 : Int;
   "2#2号电场故障" AT %I2.7 : Bool;
   "1#4号电场一次运行电压" AT %IW280 : Int;
   "1#4号电场二次运行电压" AT %IW284 : Int;
   "1#3号电场故障" AT %I1.3 : Bool;
   "2#1号电场二次运行电流" AT %IW294 : Int;
   "2#1号电场一次运行电压" AT %IW288 : Int;
   "2#1号电场二次运行电压" AT %IW292 : Int;
   "1#2号电场二次运行电压" AT %IW268 : Int;
   "1#2号电场就绪" AT %I0.5 : Bool;
   "1#2号电场备妥" AT %I0.4 : Bool;
   "1#1号电场备妥" AT %I0.0 : Bool;
   "1#1号电场故障" AT %I0.3 : Bool;
   "1#2号电场运行" AT %I0.6 : Bool;
   "1#3号电场就绪" AT %I1.1 : Bool;
   "1#4号电场备妥" AT %I1.4 : Bool;
   "1#4号电场故障" AT %I1.7 : Bool;
   "2#1号电场运行" AT %I2.2 : Bool;
   "2#2号电场就绪" AT %I2.5 : Bool;
   "2#3号电场备妥" AT %I3.0 : Bool;
   "2#3号电场就绪" AT %I3.1 : Bool;
   "2#3号电场运行" AT %I3.2 : Bool;
   "2#3号电场故障" AT %I3.3 : Bool;
   "2#4号电场备妥" AT %I3.4 : Bool;
   "2#4号电场就绪" AT %I3.5 : Bool;
   "2#4号电场运行" AT %I3.6 : Bool;
   "2#4号电场故障" AT %I3.7 : Bool;
   "1#1号电场启动" AT %Q0.0 : Bool;
   "1#1号电场停止" AT %Q0.1 : Bool;
   "1#2号电场启动" AT %Q0.2 : Bool;
   "1#2号电场停止" AT %Q0.3 : Bool;
   "1#3号电场启动" AT %Q0.4 : Bool;
   "1#3号电场停止" AT %Q0.5 : Bool;
   "1#4号电场启动" AT %Q0.6 : Bool;
   "1#4号电场停止" AT %Q0.7 : Bool;
   "2#1号电场启动" AT %Q1.0 : Bool;
   "2#1号电场停止" AT %Q1.1 : Bool;
   "2#2号电场启动" AT %Q1.2 : Bool;
   "2#2号电场停止" AT %Q1.3 : Bool;
   "2#3号电场启动" AT %Q1.4 : Bool;
   "2#3号电场停止" AT %Q1.5 : Bool;
   "2#4号电场启动" AT %Q1.6 : Bool;
   "2#4号电场停止" AT %Q1.7 : Bool;
   "1#电除尘联锁" AT %Q2.0 : Bool;
   "2#电除尘联锁" AT %Q2.1 : Bool;
   "1#1号电场控制给定" AT %QW256 : Int;
   "1#2号电场控制给定" AT %QW258 : Int;
   "1#3号电场控制给定" AT %QW260 : Int;
   "1#4号电场控制给定" AT %QW262 : Int;
   "2#1号电场控制给定" AT %QW264 : Int;
   "2#2号电场控制给定" AT %QW266 : Int;
   "2#3号电场控制给定" AT %QW268 : Int;
   "2#4号电场控制给定" AT %QW270 : Int;
   "Q2_2" AT %Q2.2 : Bool;
   "Q2_3" AT %Q2.3 : Bool;
   "Q2_4" AT %Q2.4 : Bool;
   "Q2_5" AT %Q2.5 : Bool;
   "Q2_6" AT %Q2.6 : Bool;
   "Q2_7" AT %Q2.7 : Bool;
   "Q3_0" AT %Q3.0 : Bool;
   "Q3_1" AT %Q3.1 : Bool;
   "Q3_2" AT %Q3.2 : Bool;
   "Q3_3" AT %Q3.3 : Bool;
   "Q3_4" AT %Q3.4 : Bool;
   "Q3_5" AT %Q3.5 : Bool;
   "Q3_6" AT %Q3.6 : Bool;
   "Q3_7" AT %Q3.7 : Bool;
   "Clock_Byte" AT %MB1000 : Byte;
   "Clock_10Hz" AT %M1000.0 : Bool;
   "Clock_5Hz" AT %M1000.1 : Bool;
   "Clock_2.5Hz" AT %M1000.2 : Bool;
   "Clock_2Hz" AT %M1000.3 : Bool;
   "Clock_1.25Hz" AT %M1000.4 : Bool;
   "Clock_1Hz" AT %M1000.5 : Bool;
   "Clock_0.625Hz" AT %M1000.6 : Bool;
   "Clock_0.5Hz" AT %M1000.7 : Bool;
   "Tag_1" AT %MD20 : Real;
   "Tag_2" AT %MD24 : Real;
END_VAR

VAR_GLOBAL   // PLC tag table "通讯_变量表"
   "1#除尘轴伸端U1相" AT %ID336 : Real;
   "1#除尘轴伸端V1相" AT %ID340 : Real;
   "1#除尘轴伸端W1相" AT %ID344 : Real;
   "1#除尘非轴伸端U2相" AT %ID348 : Real;
   "1#除尘非轴伸端V2相" AT %ID352 : Real;
   "1#除尘非轴伸端W2相" AT %ID356 : Real;
   "1#除尘电机前轴承温度" AT %ID360 : Real;
   "2#除尘轴伸端U1相" AT %ID432 : Real;
   "2#除尘轴伸端V1相" AT %ID436 : Real;
   "2#除尘轴伸端W1相" AT %ID440 : Real;
   "2#除尘非轴伸端U2相" AT %ID444 : Real;
   "2#除尘非轴伸端V2相" AT %ID448 : Real;
   "2#除尘非轴伸端W2相" AT %ID452 : Real;
   "2#除尘电机前轴承温度" AT %ID456 : Real;
   "1#除尘电机后轴承温度" AT %ID364 : Real;
   "1#除尘风机前轴承温度" AT %ID368 : Real;
   "1#除尘风机后轴承温度" AT %ID372 : Real;
   "2#除尘风机后轴承温度" AT %ID468 : Real;
   "2#除尘电机后轴承温度" AT %ID460 : Real;
   "2#除尘风机前轴承温度" AT %ID464 : Real;
   "QB4" AT %QB4 : Byte;
END_VAR

DATA_BLOCK "模拟量转换DB块"   // DB1
{ S7_Optimized_Access := 'FALSE' }
VERSION : 0.1
   VAR
      "1#1号电场二次运行电压" : Real := 0.0;
      "1#1号电场二次运行电流" : Real := 0.0;
      "1#2号电场二次运行电压" : Real := 0.0;
      "1#2号电场二次运行电流" : Real := 0.0;
      "1#3号电场二次运行电压" : Real := 0.0;
      "1#3号电场二次运行电流" : Real := 0.0;
      "1#4号电场二次运行电压" : Real := 0.0;
      "1#4号电场二次运行电流" : Real := 0.0;
      "2#1号电场二次运行电压" : Real := 0.0;
      "2#1号电场二次运行电流" : Real := 0.0;
      "2#2号电场二次运行电压" : Real := 0.0;
      "2#2号电场二次运行电流" : Real := 0.0;
      "2#3号电场二次运行电压" : Real := 0.0;
      "2#3号电场二次运行电流" : Real := 0.0;
      "2#4号电场二次运行电压" : Real := 0.0;
      "2#4号电场二次运行电流" : Real := 0.0;
      "1#电场热风管入口压力" : Real := 0.0;
      "1#电场热风管出口压力" : Real := 0.0;
      "2#电场热风管入口压力" : Real := 0.0;
      "2#电场热风管出口压力" : Real := 0.0;
      "1#除尘热风管进口温度" : Real := 0.0;   // -useless
      "1#除尘热风管出口温度" : Real := 0.0;   // -useless
      "2#除尘热风管进口温度" : Real;   // -useless
      "2#除尘热风管出口温度" : Real;   // -useless
      BIPOLAR : Bool;   // 单极性，始终为0
      RET_VAL : Word := WORD#16#0000;   // 错误代码
   END_VAR
BEGIN
END_DATA_BLOCK

DATA_BLOCK "百特巡检仪温度DB块"   // DB2
{ S7_Optimized_Access := 'FALSE' }